      on Press: SetTag("DB_OP.RC2", 65); SetBit("DB_OP.OP_SELMANU2")
      Visibility <- "Selec_Pleg"
      Appearance <- "DB_OP.RC2"
   Button "Botón_24" at 806,633 size 77x33; TextOff 'Retroceso'
      on Press: SetTag("DB_OP.RC2", 66); SetBit("DB_OP.OP_SELMANU2")
      Visibility <- "Selec_Pleg"
      Appearance <- "DB_OP.RC2"
   Button "Botón_25" at 889,596 size 69x33; TextOff 'Bloquear'
      on Press: SetTag("DB_OP.RC2", 20); SetBit("DB_OP.OP_SELMANU2")
      Visibility <- "Selec_Pleg"
      Appearance <- "DB_OP.RC2"
   Button "Botón_26" at 889,633 size 69x33; TextOff 'Desbloquear'
      on Press: SetTag("DB_OP.RC2", 21); SetBit("DB_OP.OP_SELMANU2")
      Visibility <- "Selec_Pleg"
      Appearance <- "DB_OP.RC2"
   Button "Botón_27" at 979,633 size 85x33; TextOff 'Bajar Prensa'
      on Press: SetTag("DB_OP.RC2", 22); SetBit("DB_OP.OP_SELMANU2")
      Visibility <- "Selec_Pleg"
      Appearance <- "DB_OP.RC2"
   Button "Botón_28" at 979,596 size 85x33; TextOff 'Subir Prensa'
      on Press: SetTag("DB_OP.RC2", 23); SetBit("DB_OP.OP_SELMANU2")
      Visibility <- "Selec_Pleg"
      Appearance <- "DB_OP.RC2"
   Button "Botón_29" at 1071,633 size 85x33; TextOff 'Bajar Ext 1'
      on Press: SetTag("DB_OP.RC2", 24); SetBit("DB_OP.OP_SELMANU2")
      Visibility <- "Selec_Pleg"
      Appearance <- "DB_OP.RC2"
   Button "Botón_30" at 1071,596 size 85x33; TextOff 'Subir Ext 1'
      on Press: SetTag("DB_OP.RC2", 25); SetBit("DB_OP.OP_SELMANU2")
      Visibility <- "Selec_Pleg"
      Appearance <- "DB_OP.RC2"
   Button "Botón_31" at 1162,633 size 85x33; TextOff 'Bajar Ext 2'
      on Press: SetTag("DB_OP.RC2", 26); SetBit("DB_OP.OP_SELMANU2")
      Visibility <- "Selec_Pleg"
      Appearance <- "DB_OP.RC2"
   Button "Botón_32" at 1162,596 size 85x33; TextOff 'Subir Ext 2'
      on Press: SetTag("DB_OP.RC2", 27); SetBit("DB_OP.OP_SELMANU2")
      Visibility <- "Selec_Pleg"
      Appearance <- "DB_OP.RC2"
   Polyline "Línea poligonal_3" at 1025,674 size 69x11
      Visibility <- "Selec_Pleg"
   TextField "Campo de texto_20" at 1097,675 size 40x18; Text 'Prensa'
      Visibility <- "Selec_Pleg"
   Polyline "Línea poligonal_4" at 1140,674 size 69x11
      Visibility <- "Selec_Pleg"
   Button "Botón_33" at 730,596 size 69x33; TextOff 'Subir'
      on Press: SetTag("DB_OP.RC2", 4); SetBit("DB_OP.OP_SELMANU2")
      Visibility <- "Selec_Pleg"
      Appearance <- "DB_OP.RC2"
   Button "Botón_34" at 730,633 size 69x33; TextOff 'Bajar'
      on Press: SetTag("DB_OP.RC2", 3); SetBit("DB_OP.OP_SELMANU2")
      Visibility <- "Selec_Pleg"
      Appearance <- "DB_OP.RC2"
   Button "Botón_35" at 806,596 size 77x33; TextOff 'Avance'
      on Press: SetTag("DB_OP.RC2", 1); SetBit("DB_OP.OP_SELMANU2")
      Visibility <- "Selec_Pleg"
      Appearance <- "DB_OP.RC2"
   Button "Botón_36" at 806,633 size 77x33; TextOff 'Retroceso'
      on Press: SetTag("DB_OP.RC2", 2); SetBit("DB_OP.OP_SELMANU2")
      Visibility <- "Selec_Pleg"
      Appearance <- "DB_OP.RC2"
   Button "Botón_37" at 889,596 size 69x33; TextOff 'Abrir'
      on Press: SetTag("DB_OP.RC2", 5); SetBit("DB_OP.OP_SELMANU2")
      Visibility <- "Selec_Pleg"
      Appearance <- "DB_OP.RC2"
   Button "Botón_38" at 889,633 size 69x33; TextOff 'Cerrar'
      on Press: SetTag("DB_OP.RC2", 6); SetBit("DB_OP.OP_SELMANU2")
      Visibility <- "Selec_Pleg"
      Appearance <- "DB_OP.RC2"
   Button "Botón_39" at 979,596 size 85x33; TextOff 'Alineación X'
      on Press: SetTag("DB_OP.RC2", 7); SetBit("DB_OP.OP_SELMANU2")
      Visibility <- "Selec_Pleg"
      Appearance <- "DB_OP.RC2"
   Button "Botón_40" at 979,633 size 85x33; TextOff 'Alineación Y'
      on Press: SetTag("DB_OP.RC2", 8); SetBit("DB_OP.OP_SELMANU2")
      Visibility <- "Selec_Pleg"
      Appearance <- "DB_OP.RC2"
   Button "Botón_41" at 1071,596 size 85x33; TextOff 'Subir Cepillos'
      on Press: SetTag("DB_OP.RC2", 9); SetBit("DB_OP.OP_SELMANU2")
      Visibility <- "Selec_Pleg"
      Appearance <- "DB_OP.RC2"
   Polyline "Línea poligonal_1" at 763,674 size 61x11
      Visibility <- "Selec_Pleg"
   TextField "Campo de texto_21" at 825,675 size 43x18; Text 'Tenaza'
      Visibility <- "Selec_Pleg"
   Polyline "Línea poligonal_2" at 873,674 size 61x11
      Visibility <- "Selec_Pleg"

screen "eProC - 10 - Estados F" 1280x770, template "Template"
   Rectangle "Rectángulo_1" at 146,344 size 393x149
      Visibility <- "STOP_RUN"
   Button "Botón_2" at 352,429 size 144x40; TextOff 'Reset'
      on Click: SetBit("PL_Reset")
      Visibility <- "STOP_RUN"
   Button "Botón_1" at 192,429 size 144x40; TextOff 'Continuar'
      on Click: SetBit("PL_Continuar")
      Visibility <- "STOP_RUN"
   TextField "Campo de texto_17" at 165,356 size 351x73; Text 'Se ha detectado un reinicio del PLC. ¿Qué desea hacer con el ciclo de la Plegadora?'
      Visibility <- "STOP_RUN"
   IOField "Champ E/S_8" at 925,320 size 99x24; Authorization "Nivel 3"; FormatPattern 999; Unit  %
      ProcessValue <- "DB_OP.PI_COD_VIT1"
   IOField "Champ E/S_4" at 926,240 size 91x29; Authorization "Nivel 2"; FormatPattern 9.9; Unit  
      ProcessValue <- "DB_OP.PI_COD_COEF"
   IOField "Champ E/S_6" at 926,260 size 91x29; Authorization "Nivel 2"; FormatPattern s9999999; Unit  mm
      ProcessValue <- "DB_OP.PI_COD_OFFSET"
   Button "Botón_6" at 779,463 size 58x33; TextOff 'Avance'
      on Press: SetTag("DB_OP.RC2", 31); SetBit("DB_OP.OP_SELMANU2")
      Visibility <- "MANU"
      Appearance <- "DB_OP.RC2"
   Button "Botón_7" at 834,463 size 58x33; TextOff 'Retroc.'
      on Press: SetTag("DB_OP.RC2", 32); SetBit("DB_OP.OP_SELMANU2")
      Visibility <- "MANU"
      Appearance <- "DB_OP.RC2"
   Button "Botón_8" at 910,463 size 58x33; TextOff 'Abrir'
      on Press: SetTag("DB_OP.RC2", 33); SetBit("DB_OP.OP_SELMANU2")
      Visibility <- "MANU"
      Appearance <- "DB_OP.RC2"
   Button "Botón_9" at 966,463 size 58x33; TextOff 'Cerrar'
      on Press: SetTag("DB_OP.RC2", 34); SetBit("DB_OP.OP_SELMANU2")
      Visibility <- "MANU"
      Appearance <- "DB_OP.RC2"
   Button "Botón_34" at 966,514 size 58x33; TextOff 'Bajar'
      on Press: SetTag("DB_OP.RC2", 40); SetBit("DB_OP.OP_SELMANU2")
      Visibility <- "MANU"
      Appearance <- "DB_OP.RC2"
   Button "Botón_35" at 909,514 size 58x33; TextOff 'Subir'
      on Press: SetTag("DB_OP.RC2", 41); SetBit("DB_OP.OP_SELMANU2")
      Visibility <- "MANU"
      Appearance <- "DB_OP.RC2"
   TextField "Campo de texto_170" at 717,678 size 17x18; Text 'F1'
   IOField "Champ E/S_162" at 732,675 size 51x25; FormatPattern s999999
      ProcessValue <- "Pinza\Pinza.PL1_1"
      Appearance <- "Pinza\Pinza.PresenciaPieza"
   IOField "Champ E/S_163" at 813,675 size 51x25; FormatPattern s999999
      ProcessValue <- "Pinza\Pinza.PL1_2"
      Appearance <- "Pinza\Pinza.PresenciaPieza"
   IOField "Champ E/S_164" at 894,675 size 51x24; FormatPattern s999999
      ProcessValue <- "Pinza\Pinza.PL2_1"
      Appearance <- "Pinza\Pinza.PresenciaPieza"
   IOField "Champ E/S_165" at 976,675 size 51x25; FormatPattern s999999
      ProcessValue <- "Pinza\Pinza.PL2_2"
      Appearance <- "Pinza\Pinza.PresenciaPieza"
   TextField "Campo de texto_171" at 797,678 size 17x18; Text 'F2'
   TextField "Campo de texto_172" at 877,678 size 17x18; Text 'F3'
   TextField "Campo de texto_173" at 959,678 size 17x18; Text 'F4'
   Button "Botón_20" at 910,576 size 58x33; TextOff 'ON'
      on Press: SetTag("DB_OP.RC2", 42); SetBit("DB_OP.OP_SELMANU2")
      Visibility <- "MANU"
      Appearance <- "DB_OP.RC2"
   Button "Botón_21" at 910,615 size 58x33; TextOff 'ON'
      on Press: SetTag("DB_OP.RC2", 46); SetBit("DB_OP.OP_SELMANU2")
      Visibility <- "MANU"
      Appearance <- "DB_OP.RC2"
   Button "Botón_22" at 966,576 size 58x33; TextOff 'OFF'
      on Press: SetTag("DB_OP.RC2", 43); SetBit("DB_OP.OP_SELMANU2")
      Visibility <- "MANU"
      Appearance <- "DB_OP.RC2"
   Button "Botón_23" at 966,615 size 58x33; TextOff 'OFF'
      on Press: SetTag("DB_OP.RC2", 47); SetBit("DB_OP.OP_SELMANU2")
      Visibility <- "MANU"
      Appearance <- "DB_OP.RC2"
   Button "Botón_28" at 786,576 size 58x33; TextOff 'ON'
      on Press: SetTag("DB_OP.RC2", 44); SetBit("DB_OP.OP_SELMANU2")
      Visibility <- "MANU"
      Appearance <- "DB_OP.RC2"
   Button "Botón_5" at 786,614 size 58x33; TextOff 'ON'
      on Press: SetTag("DB_OP.RC2", 48); SetBit("DB_OP.OP_SELMANU2")
      Visibility <- "MANU"
      Appearance <- "DB_OP.RC2"
   Button "Botón_10" at 842,576 size 58x33; TextOff 'OFF'
      on Press: SetTag("DB_OP.RC2", 45); SetBit("DB_OP.OP_SELMANU2")
      Visibility <- "MANU"
      Appearance <- "DB_OP.RC2"
   Button "Botón_31" at 842,614 size 58x33; TextOff 'OFF'
      on Press: SetTag("DB_OP.RC2", 49); SetBit("DB_OP.OP_SELMANU2")
      Visibility <- "MANU"
      Appearance <- "DB_OP.RC2"
   TextField "Template_Plantilla_Campo de texto_2" at 696,442 size 568x224; Text 'Text'
      Visibility <- "MANU"
   Circle "Círculo_2" at 78,143 size 450x450
      Appearance <- "PL_en_Ciclo"
   SymbolicIOField "Campo ES simbólico_1" at 109,310 size 387x69; TextOn '1'; TextOff '0'; TextList "Estados_F"
      ProcessValue <- "F_Estados"
   Polygon "Polígono_1" at 466,215 size 12x13
      Appearance <- "PL_en_Ciclo"
   Polygon "Polígono_2" at 520,333 size 8x12
      Appearance <- "PL_en_Ciclo"
   Polygon "Polígono_3" at 503,456 size 8x12
      Appearance <- "PL_en_Ciclo"
   Polygon "Polígono_4" at 427,543 size 14x10
      Appearance <- "PL_en_Ciclo"
   Polygon "Polígono_5" at 218,575 size 13x8
      Appearance <- "PL_en_Ciclo"
   Polygon "Polígono_6" at 124,503 size 10x13
      Appearance <- "PL_en_Ciclo"
   Polygon "Polígono_7" at 78,389 size 6x17
      Appearance <- "PL_en_Ciclo"
   Polygon "Polígono_8" at 94,269 size 7x14
      Appearance <- "PL_en_Ciclo"
   Polygon "Polígono_9" at 382,156 size 10x6
      Appearance <- "PL_en_Ciclo"
   Polygon "Polígono_10" at 162,185 size 12x9
      Appearance <- "PL_en_Ciclo"
   GraphicIOField "Campo ES gráfico_1" at 90,464 size 50x46; PictureList "Estado"
      ProcessValue <- "F_S_11"
   GraphicIOField "Campo ES gráfico_2" at 55,345 size 50x46; PictureList "Estado"
      ProcessValue <- "F_S_6"
   GraphicIOField "Campo ES gráfico_4" at 172,153 size 50x46; PictureList "Estado"
      ProcessValue <- "F_S_1"
   GraphicIOField "Campo ES gráfico_5" at 172,547 size 50x46; PictureList "Estado"
      ProcessValue <- "F_S_5"
   GraphicIOField "Campo ES gráfico_6" at 388,153 size 50x46; PictureList "Estado"
      ProcessValue <- "F_S_2"
   GraphicIOField "Campo ES gráfico_7" at 388,547 size 50x46; PictureList "Estado"
      ProcessValue <- "F_S_4"
   GraphicIOField "Campo ES gráfico_8" at 467,464 size 50x46; PictureList "Estado"
      ProcessValue <- "F_S_9"
   GraphicIOField "Campo ES gráfico_9" at 466,226 size 50x46; PictureList "Estado"
      ProcessValue <- "F_S_8"
   GraphicIOField "Campo ES gráfico_10" at 501,345 size 50x46; PictureList "Estado"
      ProcessValue <- "F_S_3"
   SymbolicIOField "Campo ES simbólico_2" at 103,359 size 403x45; TextOn '1'; TextOff '0'; TextList "Transiciones_F"
      ProcessValue <- "F_Estados"
   Line "Línea_1" at 109,126 size 0x102
      Appearance <- "PL_en_Ciclo"
   Polygon "Polígono_11" at 106,213 size 7x15
      Appearance <- "PL_en_Ciclo"
   GraphicIOField "Campo ES gráfico_11" at 84,121 size 50x46; PictureList "Estado"
      ProcessValue <- "F_S_0"
   GraphicIOField "Campo ES gráfico_3" at 86,226 size 50x46; PictureList "Estado"
      ProcessValue <- "F_S_12"
   TextField "Campo de texto_1" at 31,36 size 247x29; Text 'Máquina de estados Pinza'
   IOField "Campo ES_1" at 922,73 size 80x32; FormatPattern 9999999; Unit  mm
      ProcessValue <- "PosiciónEspera_F"
      Appearance <- "F_Req_Pos_Espera"
   TextField "Campo de texto_2" at 679,76 size 231x25; Text 'Posición de Recepción'
      Appearance <- "F_En_Pos_Espera"
   IOField "Campo ES_2" at 922,97 size 80x32; FormatPattern 9999999; Unit  mm
      ProcessValue <- "PosiciónE1H1_F"
      Appearance <- "F_Req_Pos_E1H1"
   TextField "Campo de texto_3" at 679,100 size 231x25; Text 'Posición de Esquina 1 Herramienta 1'
      Appearance <- "F_En_Pos_E1H1"
   IOField "Campo ES_3" at 922,121 size 80x32; FormatPattern 9999999; Unit  mm
      ProcessValue <- "PosiciónE1H2_F"
      Appearance <- "F_Req_Pos_E1H2"
   TextField "Campo de texto_4" at 679,124 size 231x25; Text 'Posición de Esquina 1 Herramienta 2'
      Appearance <- "F_En_Pos_E1H2"
   IOField "Campo ES_4" at 922,145 size 80x32; FormatPattern 9999999; Unit  mm
      ProcessValue <- "PosiciónE2H1_F"
      Appearance <- "F_Req_Pos_E2H1"
   TextField "Campo de texto_5" at 679,148 size 231x25; Text 'Posición de Esquina 2 Herramienta 1'
      Appearance <- "F_En_Pos_E2H1"
   IOField "Campo ES_5" at 922,169 size 80x32; FormatPattern 9999999; Unit  mm
      ProcessValue <- "PosiciónE2H2_F"
      Appearance <- "F_Req_Pos_E2H2"
   TextField "Campo de texto_6" at 679,168 size 231x25; Text 'Posición de Esquina 2 Herramienta 2'
      Appearance <- "F_En_Pos_E2H2"
   TextField "Campo de texto_9" at 679,219 size 231x25; Text 'Límite Máximo de Posición'
   IOField "Campo ES_11" at 915,216 size 88x32; FormatPattern 9999999; Unit  mm
      ProcessValue <- "PosiciónMáxima_F"
   TextField "Campo de texto_11" at 775,295 size 135x25; Text 'Posición Actual'
   IOField "Campo ES_15" at 922,291 size 128x32; FormatPattern 9999999; Unit  mm
      ProcessValue <- "PosiciónActual_F"
   TextField "Campo de texto_12" at 775,320 size 135x25; Text 'Setpoint Velocidad'
   GraphicIOField "Campo ES gráfico_12" at 276,121 size 50x46; PictureList "Estado"
      ProcessValue <- "F_S_7"
   Polygon "Polígono_12" at 262,144 size 14x5
      Appearance <- "PL_en_Ciclo"
   GraphicIOField "Campo ES gráfico_13" at 276,567 size 50x46; PictureList "Estado"
      ProcessValue <- "F_S_10"
   Polygon "Polígono_13" at 323,587 size 15x6
      Appearance <- "PL_en_Ciclo"
   IOField "Campo ES_6" at 922,193 size 80x32; FormatPattern 9999999; Unit  mm
      ProcessValue <- "PosiciónEntrega_F"
      Appearance <- "F_Req_Pos_Entrega"
   TextField "Campo de texto_8" at 679,196 size 231x25; Text 'Posición de Entrega'
      Appearance <- "F_En_Pos_Entrega"
   TextField "Campo de texto_14" at 292,131 size 16x25; Text '7'
   TextField "Campo de texto_15" at 404,163 size 16x25; Text '2'
   TextField "Campo de texto_16" at 482,236 size 16x25; Text '8'
   TextField "Campo de texto_21" at 518,355 size 16x25; Text '3'
   TextField "Campo de texto_22" at 483,474 size 16x25; Text '9'
   TextField "Campo de texto_24" at 404,557 size 16x25; Text '4'
   TextField "Campo de texto_25" at 286,577 size 30x25; Text '10'
   TextField "Campo de texto_26" at 188,557 size 19x25; Text '5'
   TextField "Campo de texto_27" at 100,474 size 30x25; Text '11'
   TextField "Campo de texto_28" at 70,355 size 15x25; Text '6'
   TextField "Campo de texto_29" at 96,236 size 31x25; Text '12'
   TextField "Campo de texto_30" at 188,163 size 16x25; Text '1'
   TextField "Campo de texto_31" at 100,131 size 16x25; Text '0'
   GraphicIOField "Campo ES gráfico_14" at 756,404 size 28x28; PictureList "CheckBox"
      ProcessValue <- "F_Tenaza_No"
   GraphicIOField "Campo ES gráfico_15" at 834,404 size 28x28; PictureList "CheckBox"
      ProcessValue <- "F_H1_No"
   GraphicIOField "Campo ES gráfico_16" at 899,404 size 28x28; PictureList "CheckBox"
      ProcessValue <- "F_H2_No"
   GraphicIOField "Campo ES gráfico_17" at 1106,401 size 28x28; PictureList "CheckBox"
      ProcessValue <- "F_Descargador_No"
   GraphicIOField "Campo ES gráfico_18" at 1195,401 size 28x28; PictureList "CheckBox"
      ProcessValue <- "F_Referencia_Menor_Descargador"
   IOField "Campo ES_7" at 1018,73 size 80x32; FormatPattern 9999999; Unit  mm
      ProcessValue <- "PosiciónEspera_F(Ant)"
   IOField "Campo ES_8" at 1018,97 size 80x32; FormatPattern 9999999; Unit  mm
      ProcessValue <- "PosiciónE1H1_F(Ant)"
   IOField "Campo ES_9" at 1018,121 size 80x32; FormatPattern 9999999; Unit  mm
      ProcessValue <- "PosiciónE1H2_F(Ant)"
   IOField "Campo ES_10" at 1018,145 size 80x32; FormatPattern 9999999; Unit  mm
      ProcessValue <- "PosiciónE2H1_F(Ant)"
   IOField "Campo ES_12" at 1018,169 size 80x32; FormatPattern 9999999; Unit  mm
      ProcessValue <- "PosiciónE2H2_F(Ant)"
   IOField "Campo ES_13" at 1018,193 size 80x32; FormatPattern 9999999; Unit  mm
      ProcessValue <- "PosiciónEntrega_F(Ant)"
   TextField "Campo de texto_34" at 249,678 size 130x18; Text 'DATOS PIEZA ACTUAL'
   TextField "Campo de texto_35" at 403,678 size 12x18; Text 'A'
   IOField "Champ E/S_24" at 414,675 size 53x25; FormatPattern 9999999
      ProcessValue <- "Pinza\Pinza.A"
      Appearance <- "Pinza\Pinza.PresenciaPieza"
   IOField "Champ E/S_25" at 483,675 size 53x25; FormatPattern 9999999
      ProcessValue <- "Pinza\Pinza.B"
      Appearance <- "Pinza\Pinza.PresenciaPieza"
   IOField "Champ E/S_26" at 554,675 size 53x24; FormatPattern 9999999
      ProcessValue <- "Pinza\Pinza.C"
      Appearance <- "Pinza\Pinza.PresenciaPieza"
   IOField "Champ E/S_27" at 629,675 size 53x25; FormatPattern 9999999
      ProcessValue <- "Pinza\Pinza.D"
      Appearance <- "Pinza\Pinza.PresenciaPieza"
   TextField "Campo de texto_36" at 472,678 size 11x18; Text 'B'
   TextField "Campo de texto_37" at 541,678 size 11x18; Text 'C'
   TextField "Campo de texto_38" at 616,678 size 12x18; Text 'D'
   TextField "Campo de texto_32" at 696,37 size 42x23; Text 'Pinza'
   TextField "Template_Plantilla_Campo de texto_4" at 696,67 size 568x3; Text 'Text'
   TextField "Template_Plantilla_Campo de texto_1" at 696,439 size 568x3; Text 'Text'
   TextField "Campo de texto_7" at 947,396 size 82x36; Text 'MOVIMIENTO SEGURO'
      Visibility <- "F_MovimientoSeguro"
      Appearance <- "F_MovimientoSeguro"
   TextField "Campo de texto_33" at 726,368 size 87x33; Text 'Tenaza Pleg. Atrás'
   TextField "Campo de texto_39" at 815,368 size 63x33; Text 'Herr. 1 OFF'
   TextField "Template_Plantilla_Campo de texto_3" at 696,359 size 568x3; Text 'Text'
   TextField "Campo de texto_43" at 882,368 size 63x33; Text 'Herr. 2 OFF'
   TextField "Campo de texto_18" at 1072,368 size 95x33; Text 'Descargador Atrás'
   TextField "Campo de texto_19" at 1160,368 size 95x33; Text 'Movimiento Corto'
   TextField "Campo de texto_10" at 719,242 size 191x25; Text 'Escalador relación mecánica'
   TextField "Campo de texto_13" at 719,262 size 191x25; Text 'Offset mecánico'
   TextField "Campo de texto_20" at 949,556 size 41x18; Text 'Martillo'
      Visibility <- "MANU"
   TextField "Campo de texto_23" at 825,556 size 35x18; Text 'Matriz'
      Visibility <- "MANU"
   TextField "Campo de texto_42" at 737,581 size 42x18; Text 'Herr. 1'
      Visibility <- "MANU"
   TextField "Campo de texto_45" at 737,622 size 42x18; Text 'Herr. 2'
      Visibility <- "MANU"
   TextField "Campo de texto_44" at 739,471 size 31x18; Text 'Pinza'
      Visibility <- "MANU"
   GraphicView "Visor de gráficos_1" at 1047,570 size 74x43; Picture "EMR2"
      Visibility <- "MANU"
   GraphicView "Visor de gráficos_2" at 1048,612 size 74x43; Picture "F1-3 EMR2"
      Visibility <- "MANU"
   GraphicView "Visor de gráficos_3" at 1152,612 size 74x43; Picture "F2-4 EMR2"
      Visibility <- "MANU"
   GraphicView "Visor de gráficos_4" at 1150,570 size 74x43; Picture "F1-3 EMR2"
      Visibility <- "MANU"
   GraphicView "Visor de gráficos_5" at 1126,590 size 12x12; Picture "outline_arrow_forward_ios_white_18dp"
      Visibility <- "MANU"
   GraphicView "Visor de gráficos_6" at 1135,590 size 12x12; Picture "outline_arrow_forward_ios_white_18dp"
      Visibility <- "MANU"
   GraphicView "Visor de gráficos_7" at 1126,632 size 12x12; Picture "outline_arrow_forward_ios_white_18dp"
      Visibility <- "MANU"
   GraphicView "Visor de gráficos_8" at 1135,632 size 12x12; Picture "outline_arrow_forward_ios_white_18dp"
      Visibility <- "MANU"
   TextField "Campo de texto_40" at 740,522 size 134x18; Text 'Bloque de Herramientas'
      Visibility <- "MANU"
   Button "Botón_42" at 48,625 size 40x40; TextOff 'Vista Condiciones'; PictureOff "Gráfico_7"
      on Click: ActivateScreen("eProC - 10 - Estados F_HW", 0)
   Button "Botón_11" at 1224,27 size 40x37; TextOff 'Vista Condiciones'; PictureOff "Tool"; Authorization "Nivel 3"
      on Click: ActivateScreen("eProC - 11 Referencias F-PL", 0)

screen "eProC - 10 - Estados F_HW" 1280x770, template "Template"
   GraphicIOField "Campo ES gráfico_6" at 554,292 size 718x282; PictureList "Grupo 3 - Pinza1"
      ProcessValue <- "Alarma_Pinza"
   Polygon "Polígono_2" at 281,432 size 517x163
      Visibility <- "Pinza\Pinza.PresenciaPieza"
   Circle "Cercle_16" at 798,434 size 10x10
      Appearance <- "29S4"
   TextField "Campo de texto_29" at 910,349 size 114x18; Text '29S4 - Pinza Abierta'
   TextField "Campo de texto_30" at 894,313 size 116x18; Text '29S5 - Pinza Cerrada'
   Circle "Cercle_17" at 798,418 size 10x10
      Appearance <- "29S5"
   GraphicIOField "Campo ES gráfico_8" at 192,179 size 289x268; PictureList "Formador"
      ProcessValue <- "Alarma_Formador"
   Circle "Cercle_6" at 331,217 size 10x10
      Appearance <- "28S5"
   Circle "Cercle_7" at 331,246 size 10x10
      Appearance <- "28S6"
   TextField "Campo de texto_3" at 54,201 size 180x18; Text '28S5 - Herramientas Bloqueadas'
   TextField "Campo de texto_5" at 36,229 size 200x18; Text '28S6 - Herramientas Desbloqueadas'
   Circle "Cercle_8" at 406,291 size 10x10
      Appearance <- "28S3"
   Circle "Cercle_9" at 418,306 size 10x10
      Appearance <- "28S4"
   Circle "Cercle_10" at 460,360 size 10x10
      Appearance <- "28S1"
   Circle "Cercle_1" at 437,332 size 10x10
      Appearance <- "28S2"
   Circle "Cercle_0" at 371,397 size 10x10
      Appearance <- "27S5"
   Circle "Cercle_2" at 348,367 size 10x10
      Appearance <- "27S6"
   Circle "Cercle_18" at 313,326 size 10x10
      Appearance <- "27S7"
   Circle "Cercle_19" at 326,344 size 10x10
      Appearance <- "27S8"
   TextField "Campo de texto_10" at 488,240 size 146x18; Text '28S3 - Herr. 2 Matriz OFF'
   TextField "Campo de texto_15" at 496,267 size 142x18; Text '28S4 - Herr. 2 Matriz ON'
   TextField "Campo de texto_16" at 522,323 size 152x18; Text '28S1 - Herr. 2 Martillo OFF'
   TextField "Campo de texto_17" at 506,295 size 148x18; Text '28S2 - Herr. 2 Martillo ON'
   TextField "Campo de texto_11" at 44,381 size 146x18; Text '27S7 - Herr. 1 Matriz OFF'
   TextField "Campo de texto_19" at 46,411 size 142x18; Text '27S8 - Herr. 1 Matriz ON'
   TextField "Campo de texto_20" at 73,488 size 152x18; Text '27S5 - Herr. 1 Martillo OFF'
   TextField "Campo de texto_21" at 58,452 size 148x18; Text '27S6 - Herr. 1 Martillo ON'
   Button "Botón_42" at 48,625 size 40x40; TextOff 'Vista Condiciones'; PictureOff "Gráfico_6"
      on Click: ActivateScreen("eProC - 10 - Estados F", 0)
   TextField "Campo de texto_1" at 804,90 size 41x18; Text 'Martillo'
      Visibility <- "MANU"
   TextField "Campo de texto_23" at 680,90 size 35x18; Text 'Matriz'
      Visibility <- "MANU"
   TextField "Campo de texto_42" at 592,115 size 42x18; Text 'Herr. 1'
      Visibility <- "MANU"
   TextField "Campo de texto_45" at 592,156 size 42x18; Text 'Herr. 2'
      Visibility <- "MANU"
   TextField "Campo de texto_44" at 732,638 size 31x18; Text 'Pinza'
      Visibility <- "MANU"
   GraphicView "Visor de gráficos_1" at 904,108 size 74x43; Picture "EMR2"
      Visibility <- "MANU"
   GraphicView "Visor de gráficos_2" at 905,150 size 74x43; Picture "F1-3 EMR2"
      Visibility <- "MANU"
   GraphicView "Visor de gráficos_3" at 1009,150 size 74x43; Picture "F2-4 EMR2"
      Visibility <- "MANU"
   GraphicView "Visor de gráficos_4" at 1007,108 size 74x43; Picture "F1-3 EMR2"
      Visibility <- "MANU"
   GraphicView "Visor de gráficos_5" at 983,128 size 12x12; Picture "outline_arrow_forward_ios_white_18dp"
      Visibility <- "MANU"
   GraphicView "Visor de gráficos_6" at 992,128 size 12x12; Picture "outline_arrow_forward_ios_white_18dp"
      Visibility <- "MANU"
   GraphicView "Visor de gráficos_7" at 983,170 size 12x12; Picture "outline_arrow_forward_ios_white_18dp"
      Visibility <- "MANU"
   GraphicView "Visor de gráficos_8" at 992,170 size 12x12; Picture "outline_arrow_forward_ios_white_18dp"
      Visibility <- "MANU"
   TextField "Campo de texto_40" at 270,118 size 134x18; Text 'Bloque de Herramientas'
      Visibility <- "MANU"
   TextField "Campo de texto_12" at 460,410 size 81x18; Text 'Herramienta 2'
   TextField "Campo de texto_13" at 366,434 size 81x18; Text 'Herramienta 1'
   Button "Botón_6" at 772,630 size 58x33; TextOff 'Avance'
      on Press: SetTag("DB_OP.RC2", 31); SetBit("DB_OP.OP_SELMANU2")
      Visibility <- "MANU"
      Appearance <- "DB_OP.RC2"
   Button "Botón_7" at 827,630 size 58x33; TextOff 'Retroc.'
      on Press: SetTag("DB_OP.RC2", 32); SetBit("DB_OP.OP_SELMANU2")
      Visibility <- "MANU"
      Appearance <- "DB_OP.RC2"
   Button "Botón_8" at 903,630 size 58x33; TextOff 'Abrir'
      on Press: SetTag("DB_OP.RC2", 33); SetBit("DB_OP.OP_SELMANU2")
      Visibility <- "MANU"
      Appearance <- "DB_OP.RC2"
   Button "Botón_9" at 959,630 size 58x33; TextOff 'Cerrar'
      on Press: SetTag("DB_OP.RC2", 34); SetBit("DB_OP.OP_SELMANU2")
      Visibility <- "MANU"
      Appearance <- "DB_OP.RC2"
   Button "Botón_34" at 496,110 size 58x33; TextOff 'Bajar'
      on Press: SetTag("DB_OP.RC2", 40); SetBit("DB_OP.OP_SELMANU2")
      Visibility <- "MANU"
      Appearance <- "DB_OP.RC2"
   Button "Botón_35" at 439,110 size 58x33; TextOff 'Subir'
      on Press: SetTag("DB_OP.RC2", 41); SetBit("DB_OP.OP_SELMANU2")
      Visibility <- "MANU"
      Appearance <- "DB_OP.RC2"
   Button "Botón_20" at 765,110 size 58x33; TextOff 'ON'
      on Press: SetTag("DB_OP.RC2", 42); SetBit("DB_OP.OP_SELMANU2")
      Visibility <- "MANU"
      Appearance <- "DB_OP.RC2"
   Button "Botón_21" at 765,149 size 58x33; TextOff 'ON'
      on Press: SetTag("DB_OP.RC2", 46); SetBit("DB_OP.OP_SELMANU2")
      Visibility <- "MANU"
      Appearance <- "DB_OP.RC2"
   Button "Botón_22" at 821,110 size 58x33; TextOff 'OFF'
      on Press: SetTag("DB_OP.RC2", 43); SetBit("DB_OP.OP_SELMANU2")
      Visibility <- "MANU"
      Appearance <- "DB_OP.RC2"
   Button "Botón_23" at 821,149 size 58x33; TextOff 'OFF'
      on Press: SetTag("DB_OP.RC2", 47); SetBit("DB_OP.OP_SELMANU2")
      Visibility <- "MANU"
      Appearance <- "DB_OP.RC2"
   Button "Botón_28" at 641,110 size 58x33; TextOff 'ON'
      on Press: SetTag("DB_OP.RC2", 44); SetBit("DB_OP.OP_SELMANU2")
      Visibility <- "MANU"
      Appearance <- "DB_OP.RC2"
   Button "Botón_5" at 641,148 size 58x33; TextOff 'ON'
      on Press: SetTag("DB_OP.RC2", 48); SetBit("DB_OP.OP_SELMANU2")
      Visibility <- "MANU"
      Appearance <- "DB_OP.RC2"
   Button "Botón_10" at 697,110 size 58x33; TextOff 'OFF'
      on Press: SetTag("DB_OP.RC2", 45); SetBit("DB_OP.OP_SELMANU2")
      Visibility <- "MANU"
      Appearance <- "DB_OP.RC2"
   Button "Botón_31" at 697,148 size 58x33; TextOff 'OFF'
      on Press: SetTag("DB_OP.RC2", 49); SetBit("DB_OP.OP_SELMANU2")
      Visibility <- "MANU"
      Appearance <- "DB_OP.RC2"

screen "eProC - 11 Referencias F-PL" 1280x770, template "Template"
   GraphicView "Visor de gráficos_1" at 134,72 size 979x505; Picture "Referencias"
   IOField "Champ E/S" at 340,310 size 80x27; Authorization "Nivel 2"; FormatPattern 9999999
      ProcessValue <- "Distancia_entre_Herramienta1_y_Pos0_F"
   IOField "Champ E/S_0" at 540,342 size 80x26; Authorization "Nivel 2"; FormatPattern 9999999
      ProcessValue <- "Distancia_entre_Pos0_y_Tenaza_F"
   TextField "Campo de texto_1" at 334,240 size 90x68; Text 'Distancia de Herramienta 1 a posición 0mm Pinza'
   TextField "Campo de texto_3" at 526,300 size 126x36; Text 'Distancia 0mm Pinza a Tenaza Plegadora'
   IOField "Champ E/S_2" at 552,526 size 80x26; Authorization "Nivel 2"; FormatPattern 9999999
      ProcessValue <- "Distancia_entre_Pos0_y_Descargador_F"
   TextField "Campo de texto_6" at 505,553 size 176x36; Text 'Distancia posición 0mm Pinza al Descargador'
   IOField "Champ E/S_3" at 235,566 size 80x27; Authorization "Nivel 2"; FormatPattern 9999999
      ProcessValue <- "Distancia_entre_Herramientas_F"
   TextField "Campo de texto_7" at 230,594 size 93x36; Text 'Distancia entre Herramientas'
   IOField "Champ E/S_4" at 592,610 size 80x26; Authorization "Nivel 2"; FormatPattern s9999999999
      ProcessValue <- "PosiciónMáxima_F"
   TextField "Campo de texto_8" at 587,636 size 93x36; Text 'Distancia Avance Máximo'
   IOField "Champ E/S_1" at 907,300 size 80x26; Authorization "Nivel 2"; FormatPattern 9999999
      ProcessValue <- "Distancia_entre_Pleg_Alin_PL"
   TextField "Campo de texto_2" at 861,330 size 196x20; Text 'Distancia de Plegador a Alineador'
   Switch "Interruptor_1" at 209,115 size 125x80; CaptionText 'Habilitar reglas'; TextOff 'NO'; TextOn 'SI'
      ProcessValue <- "HabilitarReglasBaluff"

VB script "Script_1"
   'NOTE : Appuyez sur <Ctrl><Espacement> pour lancer le script et afficher le large éventail de fonctions.
   'Ecrivez vos scripts en utilisant les fonctions système ou le modèle d'objet. Vous pouvez facilement accéder au
   'système via l'objet runtime IHM. Pour sélectionner rapidement une référence objet
   'vous pouvez appuyer sur <Alt><Flèche droite>. Vous pouvez créer des scripts complexes en ayant recours au
   'langage de programmation VBScript et accéder directement aux variables via le nom, par ex. tag = 5.
*)